
   REGION "BUTTON SELECTION BUTTONS"
       FOR #i := 0 TO "BUTTON_COUNT" DO
           #t_interface.buttons[#i].animate := "Bool.Animate"(true_color := "GREEN_LIGHT_BACKGROUND",
                                                              false_color := "GRAY_BACKGROUND",
                                                              evaluation_signal := #interface.buttons[#i].actuate);
           #t_interface.buttons[#i].enable := TRUE;
           #t_interface.buttons[#i].visible := TRUE;
           IF #selected.btns[#i] THEN
               #t_interface.buttons[#i].animate := "BLUE_LIGHT_BACKGROUND";
           END_IF;
       END_FOR;
   END_REGION


   REGION "DRAW"
       #interface := #t_interface;
   END_REGION
END_FUNCTION

FUNCTION "Pop Up: Select Buttons: Pulse Ints to Bools" : Void   // FC118, SCL
{ S7_Optimized_Access := 'TRUE' }
VERSION : 0.1
   VAR_INPUT
      pulses_as_ints : Array[0.."BUTTON_COUNT"] of Int;
   END_VAR
   VAR_OUTPUT
      pulses_as_bools : Array[0.."BUTTON_COUNT"] of Bool;
   END_VAR
   VAR_TEMP
      i : Int;
      ret : Array[0.."BUTTON_COUNT"] of Bool;
   END_VAR
BEGIN
   REGION "MAP TO BOOLS"
       FOR #i := 0 TO "BUTTON_COUNT" DO
           #ret[#i] := #pulses_as_ints[#i].%X0;
       END_FOR;
   END_REGION

   REGION "RETURN"
       #pulses_as_bools := #ret;
   END_REGION
END_FUNCTION

// folder: Display: Warehouse/Pop Ups/Select Station

FUNCTION_BLOCK "Pop Up: Select Stations"   // FB21, SCL
{ S7_Optimized_Access := 'TRUE' }
VERSION : 0.1
   VAR_INPUT
      all_stations : "Station: All Stations";
      saved_WIPs : "Recipe: HMI Stations Saved Wips";
   END_VAR
   VAR_IN_OUT
      interface : "Select Station";
      meta_data : "Setting Meta Data";
   END_VAR
   VAR
      "inst Patch for Table Nav in Select Station Popup" : "Patch for Table Nav in Select Station Popup";
      "inst Select Station Button Pulses" : "Pulses: Button Collection";
      "inst Selection Change" : "Selected_Stations.Selection_Change";
      "inst Table Nav" : "Table Nav";
      vis_stns_as_dint : Array[0.."_SELECT_STATION_BUTTON_COUNT"] of DInt;
      visable_stns : Array[0.."_SELECT_STATION_BUTTON_COUNT"] of Int;
   END_VAR
   VAR_TEMP
      actuations_as_ints : Array[0.."_SELECT_STATION_BUTTON_COUNT"] of Int;
      actuation_pulses : Array[0.."_SELECT_STATION_BUTTON_COUNT"] of Bool;
      actuation_pulses_as_int : Array[0.."_SELECT_STATION_BUTTON_COUNT"] of Int;
      blank_station : "Station: Single Station";
      i : Int;
      nav_pulses : Int;
      p_stn : DInt;
      selectable_stns_as_dint : Array[0.."STATION_COUNT"] of DInt;
      t_selection_change : "Station Selection Change";
   END_VAR
   // visable_stns[0] := 0;
   // visable_stns[1] := 1;
   // visable_stns[2] := 2;
   // visable_stns[3] := 3;
   // visable_stns[4] := 4;
   // visable_stns[5] := 5;
   // visable_stns[6] := 6;
   // visable_stns[7] := 7;
   // visable_stns[8] := 8;
   // visable_stns[9] := 9;
   // visable_stns[10] := 10;
   // visable_stns[11] := 11;
BEGIN
   REGION "ANIMATIONS"
       "Pop Up: Select Stations: Animations"(all_stations := #all_stations,
                                             meta_data := #meta_data,
                                             visable_stns := #visable_stns,
                                             interface := #interface);
   END_REGION


   REGION "CLEAR SELECTION CHANGE"
       #meta_data.station_selection_change := #t_selection_change;
   END_REGION


   REGION "SELECT STATION BUTTON PULSES"
       "Pop Up: Map Select Button Actuations"(screen_elements := #interface.stn_select_btns,
                                              actuations_as_ints := #actuations_as_ints);
       #"inst Select Station Button Pulses"(btns := #actuations_as_ints,
                                            pulses := #actuation_pulses_as_int);
       "Pop Up: Select Stations: Pulse Ints to Bools"(pulses_as_ints := #actuation_pulses_as_int,
                                                      pulses_as_bools => #actuation_pulses);
   END_REGION


   REGION "PERFORM STATION SELECTION"
       FOR #i := 0 TO "_SELECT_STATION_BUTTON_COUNT" DO
           IF #visable_stns[#i] <> -1 THEN
               "Toggle"(pulse := #actuation_pulses[#i],
                        state := #meta_data.selected_stations.stns[#visable_stns[#i]]);
           END_IF;
       END_FOR;
       #meta_data.selected_stations.count := "Count Selected Stations"(#meta_data.selected_stations.stns);
   END_REGION


   REGION "SCAN FOR CHANGE TO STATION SELECTION"
       #"inst Selection Change"(selected_stns := #meta_data.#selected_stations,
                                station_change => #meta_data.station_selection_change);
   END_REGION


   REGION "BUILD SELECTABLE STATION LIST"
       IF #meta_data.station_selection_change.selection_change OR "FirstScan" THEN
           "Pop Up: Select Stations: Build Selectable Station List"(saved_wips := #saved_WIPs,
                                                                    all_stations := #all_stations,
                                                                    meta_data := #meta_data);
       END_IF;
   END_REGION


   REGION "TABLE NAV"

       // when there are more selectable stations than buttons
       IF #meta_data.selectable_stations.count > "_SELECT_STATION_BUTTON_COUNT" THEN
           #"inst Table Nav"(first_null_index := #meta_data.selectable_stations.count,
                             tblData := #selectable_stns_as_dint,
                             tblDisp := #vis_stns_as_dint,
                             tableNav := #interface.nav_bar.plc,
                             rowIndices := #vis_stns_as_dint);
           // patch for table nav to work with selectable stations
           #"inst Patch for Table Nav in Select Station Popup"(nav_bar := #interface.nav_bar.plc,
                                                               meta_data := #meta_data,
                                                               vis_stns_as_dint := #vis_stns_as_dint,
                                                               visable_stns := #visable_stns);
       END_IF;

       // when there are fewer selectable stations than buttons
       IF #meta_data.selectable_stations.count <= "_SELECT_STATION_BUTTON_COUNT" + 1 THEN
           IF #meta_data.station_selection_change.selection_change THEN
               "Array.Int.Fill"(value:="NULL_TOKEN",
                                int_array := #visable_stns);
               FOR #i := 0 TO #meta_data.selectable_stations.count - 1 DO
                   #visable_stns[#i] := #meta_data.selectable_stations.stns[#i];
               END_FOR;
           END_IF;
       END_IF;


   END_REGION
END_FUNCTION_BLOCK

FUNCTION_BLOCK "Selected_Stations.Selection_Change"   // FB23, SCL
{ S7_Optimized_Access := 'TRUE' }
VERSION : 0.1
   VAR_INPUT
      selected_stns : "Selected Stations";
   END_VAR
   VAR_OUTPUT
      station_change : "Station Selection Change";
   END_VAR
   VAR
      old : Struct
         selected_stns : "Selected Stations";
      END_STRUCT;
   END_VAR
   VAR_TEMP
      i : Int;
      ret : "Station Selection Change";
   END_VAR
BEGIN
   REGION "SCAN FOR CHANGE"
       FOR #i := 0 TO "STATION_COUNT" DO
           IF #selected_stns.stns[#i] <> #old.selected_stns.stns[#i] THEN
               #ret.selection_change := TRUE;
               #ret.station_index := #i;
               IF #selected_stns.stns[#i] AND NOT #old.selected_stns.stns[#i] THEN
                   #ret.rising := TRUE;
                   #ret.falling := FALSE;
               END_IF;
               IF NOT #selected_stns.stns[#i] AND #old.selected_stns.stns[#i] THEN
                   #ret.rising := FALSE;
                   #ret.falling := TRUE;
               END_IF;
               EXIT;
           END_IF;
       END_FOR;
   END_REGION


   REGION "SAVE TO OLD"
       #old.selected_stns := #selected_stns;
   END_REGION


   REGION "RETURN"
       #station_change.falling := #ret.falling;
       #station_change.rising := #ret.rising;
       #station_change.selection_change := #ret.selection_change;
       #station_change.station_index := #ret.station_index;
   END_REGION
END_FUNCTION_BLOCK

FUNCTION_BLOCK "Patch for Table Nav in Select Station Popup"   // FB24, SCL
{ S7_Optimized_Access := 'TRUE' }
VERSION : 0.1
   VAR_INPUT
      nav_bar : "Nav Bar Data: PLC";
      meta_data : "Setting Meta Data";
   END_VAR
   VAR_IN_OUT
      vis_stns_as_dint : Array[0.."_SELECT_STATION_BUTTON_COUNT"] of DInt;
      visable_stns : Array[0.."_SELECT_STATION_BUTTON_COUNT"] of Int;
   END_VAR
   VAR
      old_nav : "Nav Bar Data: PLC";
   END_VAR
   VAR_TEMP
      first_row : Int;
      i : Int;
      nav_pulse : Bool;
      p_visable_row : Int;
      search_term : Int;
      t_visable_stns : Array[0.."_SELECT_STATION_BUTTON_COUNT"] of Int;
   END_VAR
BEGIN
   REGION "PULSE FROM ANY NAV BUTTON"
       IF NOT #old_nav.top.actuate AND #nav_bar.top.actuate THEN
           #nav_pulse := TRUE;
       END_IF;
       IF NOT #old_nav.pageUp.actuate AND #nav_bar.pageUp.actuate THEN
           #nav_pulse := TRUE;
       END_IF;
       IF NOT #old_nav.lineUp.actuate AND #nav_bar.lineUp.actuate THEN
           #nav_pulse := TRUE;
       END_IF;
       IF NOT #old_nav.lineDown.actuate AND #nav_bar.lineDown.actuate THEN
           #nav_pulse := TRUE;
       END_IF;
       IF NOT #old_nav.pageDown.actuate AND #nav_bar.pageDown.actuate THEN
           #nav_pulse := TRUE;
       END_IF;
       IF NOT #old_nav.bottom.actuate AND #nav_bar.bottom.actuate THEN
           #nav_pulse := TRUE;
       END_IF;
   END_REGION



   REGION "REMAP VISIBLE STATIONS BASED ON SELECTABLE STATIONS"

       REGION "NAV REMAP"
           IF #nav_pulse THEN
               FOR #i := 0 TO "_SELECT_STATION_BUTTON_COUNT" DO
                   #t_visable_stns[#i] := #meta_data.selectable_stations.stns[DINT_TO_INT(#vis_stns_as_dint[#i])];
                   #vis_stns_as_dint[#i] := #t_visable_stns[#i];
               END_FOR;
               #visable_stns := #t_visable_stns;
           END_IF;
       END_REGION

       REGION "SELECTION REMAP"
           IF #meta_data.station_selection_change.selection_change THEN
               #search_term := #visable_stns[0];
               #first_row := "Array.Int.Search"(array_of_int := #meta_data.selectable_stations.stns,
                                                 search_term := #search_term);
               WHILE #first_row = "NULL_TOKEN" DO
                   #search_term -= 1;
                   IF #search_term < 0 THEN
                       #search_term := 0;
                       EXIT;
                   END_IF;
                   #first_row := "Array.Int.Search"(array_of_int := #meta_data.selectable_stations.stns,
                                                     search_term := #search_term);
               END_WHILE;
               // direct write access required to keep collapsed or uncollapsed
               // format after nav button press
               "EMP IDB"."inst Pop Up: Select Station"."inst Table Nav".r1 := #first_row;
               FOR #i := 0 TO "_SELECT_STATION_BUTTON_COUNT" DO
                   #p_visable_row := #first_row + #i;
                   IF #p_visable_row >= #meta_data.selectable_stations.count THEN
                       #p_visable_row -= #meta_data.selectable_stations.count;
                   END_IF;
                   #t_visable_stns[#i] := #meta_data.selectable_stations.stns[#p_visable_row];
                   #vis_stns_as_dint[#i] := #t_visable_stns[#i];
               END_FOR;
               #visable_stns := #t_visable_stns;
           END_IF;
       END_REGION
   (*    
       IF #meta_data.selection_change.selection_change THEN

           REGION "COPY TO LOCAL"
               FOR #i := 0 TO "slct_stn_btn_count" DO
                   #t_visable_stns[#i] := DINT_TO_INT(#vis_stns_as_dint[#i]);
               END_FOR;
           END_REGION



           IF #meta_data.selection_change.falling AND #meta_data.selected_stations.count = 0 THEN
               #first_row := DINT_TO_INT(#vis_stns_as_dint[0]);
               FOR #i := 0 TO "slct_stn_btn_count" DO
                   #t_visable_stns[#i] := #first_row + #i;
                   IF #t_visable_stns[#i] > "stnCount" THEN
                       #t_visable_stns[#i] -= "stnCount" + 1;
                   END_IF;
               END_FOR;
           END_IF;

           IF #meta_data.selection_change.selection_change AND #meta_data.selected_stations.count <> 0 THEN
               FOR #i := 0 TO "slct_stn_btn_count" DO
                   IF DINT_TO_INT(#vis_stns_as_dint[#i]) > #meta_data.selectable_stations.count - 1 THEN
                       #t_visable_stns[#i] := DINT_TO_INT(#vis_stns_as_dint[#i]) - #meta_data.selectable_stations.count;
                   END_IF;
                   IF DINT_TO_INT(#vis_stns_as_dint[#i]) <= #meta_data.selectable_stations.count - 1 THEN

                   END_IF;
               END_FOR;
           END_IF;


           REGION "RETURN"
               FOR #i := 0 TO "slct_stn_btn_count" DO
                   #vis_stns_as_dint[#i] := INT_TO_DINT(#t_visable_stns[#i]);
               END_FOR;
               #visable_stns := #t_visable_stns;
           END_REGION


       END_IF;
   *)    

   END_REGION


   REGION "SAVE FOR CHANGE DETECTION"
       #old_nav := #nav_bar;
   END_REGION
END_FUNCTION_BLOCK

FUNCTION "Populate Station Name" : WString   // FC100, SCL
{ S7_Optimized_Access := 'TRUE' }
VERSION : 0.1
   VAR_INPUT
      lines : Int;
      stn : "Station: Single Station";
   END_VAR
   VAR_TEMP
      ret : WString;
      dz : WString;
   END_VAR
   VAR CONSTANT
      line_feed : WString := WSTRING#'$L';
   END_VAR
BEGIN
   REGION "FORMAT STRING"
       #dz := "Strip Sign"(USINT_TO_WSTRING(#stn.id.dropZone));
       #dz := "Add Leading"("Leading Character" := wchar#'0',
                            "Desired Length" := 2,
                            "String" := #dz);
   END_REGION

   REGION "ONE LINE"
       IF #lines = 1 THEN
           #ret := CONCAT_WSTRING(IN1 := #stn.id.lineName,
                                  IN2 := #dz);
       END_IF;
   END_REGION


   REGION "MORE THAN ONE LINE"
       IF #lines > 1 THEN
           #ret := CONCAT_WSTRING(IN1 := #stn.id.lineName,
                                  IN2 := #line_feed,
                                  IN3 := #dz);
       END_IF;
   END_REGION


   REGION "INVALID ENTRY"
       IF #lines < 1 THEN
           #ret := WString#'invalid line count';
       END_IF;
   END_REGION


   #"Populate Station Name" := #ret;
END_FUNCTION

FUNCTION "Pop Up: Select Stations: Map Select Button Acutations" : Void   // FC101, SCL
{ S7_Optimized_Access := 'TRUE' }
VERSION : 0.1
   VAR_INPUT
      select_btns : Array[0.."_SELECT_STATION_BUTTON_COUNT"] of "Push Button Data";
   END_VAR
   VAR_OUTPUT
      btn_actuations : Array[0.."_SELECT_STATION_BUTTON_COUNT"] of Int;
   END_VAR
   VAR_TEMP
      i : Int;
      ret : Array[0.."_SELECT_STATION_BUTTON_COUNT"] of Int;
   END_VAR
BEGIN
   REGION "MAP ACTUATIONS"
       FOR #i := 0 TO "_SELECT_STATION_BUTTON_COUNT" DO
           IF #select_btns[#i].actuate THEN
               #ret[#i] := 1;
           END_IF;
       END_FOR;
   END_REGION


   REGION "RETURN"
       #btn_actuations := #ret;
   END_REGION
END_FUNCTION

FUNCTION "Pop Up: Select Stations: Pulse Ints to Bools" : Void   // FC102, SCL
{ S7_Optimized_Access := 'TRUE' }
VERSION : 0.1
   VAR_INPUT
      pulses_as_ints : Array[0.."_SELECT_STATION_BUTTON_COUNT"] of Int;
   END_VAR
   VAR_OUTPUT
      pulses_as_bools : Array[0.."_SELECT_STATION_BUTTON_COUNT"] of Bool;
   END_VAR
   VAR_TEMP
      i : Int;
      ret : Array[0.."_SELECT_STATION_BUTTON_COUNT"] of Bool;
   END_VAR
BEGIN
   REGION "MAP TO BOOLS"
       FOR #i := 0 TO "_SELECT_STATION_BUTTON_COUNT" DO
           #ret[#i] := #pulses_as_ints[#i].%X0;
       END_FOR;
   END_REGION

   REGION "RETURN"
       #pulses_as_bools := #ret;
   END_REGION
END_FUNCTION

FUNCTION "Pop Up: Select Stations: Build Selectable Station List" : Void   // FC104, SCL
{ S7_Optimized_Access := 'TRUE' }
VERSION : 0.1
   VAR_INPUT
      saved_wips : "Recipe: HMI Stations Saved Wips";
      all_stations : "Station: All Stations";
   END_VAR
   VAR_IN_OUT
      meta_data : "Setting Meta Data";
   END_VAR
   VAR_TEMP
      eval_station_is_hmi : Bool;
      blank_stn : "Station: Single Station";
      i : Int;
      states : "Selectable Station States";
      md : "Setting Meta Data";
   END_VAR
   VAR CONSTANT
      initialize : String := 'initialize';
      all : String := 'all';
      non_hmi : String := 'non_hmi';
      hmi : String := 'hmi';
   END_VAR
BEGIN
   REGION "NOTES"
       (*
       The UDT containing all stations is too large to be instantiated in temp
       memory for this function. This is why you will see an initialization loop
       instead of a temp variable that gets returned later.
       *)
   END_REGION


   REGION "FOR ANY STATE"

       REGION "COPY TO LOCAL"
           #md := #meta_data;
       END_REGION

       REGION "SELECTED STATION IS HMI"
           IF #md.station_selection_change.rising THEN
               #eval_station_is_hmi := "Station.Is_HMI_Station"(#all_stations.stn[#md.station_selection_change.station_index]);
           END_IF;
           IF #md.station_selection_change.falling AND #md.selected_stations.count = 1 THEN
               #eval_station_is_hmi := "Station.Is_HMI_Station"(#all_stations.stn["Get First Selected Station"(#md.selected_stations.stns)]);
           END_IF;
       END_REGION

   END_REGION


   REGION "SET STATE"

       REGION "ALL"
           // on first scan
           IF "FirstScan" THEN
               #states := "Set Selectable Station States"(#all);
               GOTO EVAL;
           END_IF;
           // on selection change where last selected station is de-selected
           IF #md.station_selection_change.falling AND #md.selected_stations.count = 0 THEN
               #states := "Set Selectable Station States"(#all);
               GOTO EVAL;
           END_IF;
       END_REGION

       REGION "NON HMI"
           // when no stations are selected and a non-hmi station is selected
           IF #md.station_selection_change.selection_change (*AND #selected_stn_count = 1*) THEN
               IF NOT #eval_station_is_hmi THEN
                   #states := "Set Selectable Station States"(#non_hmi);
                   GOTO EVAL;
               END_IF;
           END_IF;
       END_REGION

       REGION "HMI"
           // when no stations are selected and an hmi station is selected
           IF #md.station_selection_change.selection_change (*AND #selected_stn_count = 1*) THEN
               IF #eval_station_is_hmi THEN
                   #states := "Set Selectable Station States"(#hmi);
                   GOTO EVAL;
               END_IF;
           END_IF;
       END_REGION

   END_REGION


   REGION "STATE LOGIC"
   EVAL:

       REGION "ALL"
           IF #states.all THEN
               "Array.Int.Fill"(value:="NULL_TOKEN",
                                int_array := #md.selectable_stations.stns);
               FOR #i := 0 TO "STATION_COUNT" DO
                   #md.selectable_stations.stns[#i] := #i;
               END_FOR;
               #md.selectable_stations.count := "STATION_COUNT" + 1;
               GOTO RTRN;
           END_IF;
       END_REGION


       REGION "NON-HMI"
           IF #states.non_hmi THEN
               "Array.Int.Fill"(value:="NULL_TOKEN",
                                int_array := #md.selectable_stations.stns);
               #md.selectable_stations := "Pop Up: Select Stations: Build Non-HMI List"(#all_stations);
               GOTO RTRN;
           END_IF;
       END_REGION


       REGION "HMI"
           IF #states.hmi THEN
               "Array.Int.Fill"(value:="NULL_TOKEN",
                                int_array := #md.selectable_stations.stns);
               #md.selectable_stations := "Pop Up: Select Stations: Build HMI List"(saved_wips := #saved_wips,
                                                                                    meta_data := #md);
               GOTO RTRN;
           END_IF;
       END_REGION

   END_REGION


   REGION "RETURN"
   RTRN:
       #meta_data := #md;
   END_REGION
END_FUNCTION

FUNCTION "Set Selectable Station States" : "Selectable Station States"   // FC107, SCL
{ S7_Optimized_Access := 'TRUE' }
VERSION : 0.1
   VAR_INPUT
      desired_state : String;
   END_VAR
   VAR_TEMP
      ret : "Selectable Station States";
   END_VAR
   VAR CONSTANT
      initialize : String := 'initialize';
      all : String := 'all';
      non_hmi : String := 'non_hmi';
      hmi : String := 'hmi';
   END_VAR
BEGIN
   REGION "SET ALL"
       IF #desired_state = #all THEN
           #ret.all := TRUE;
       END_IF;
   END_REGION


   REGION "SET NON_HMI"    
       IF #desired_state = #non_hmi THEN
           #ret.non_hmi := TRUE;
       END_IF;
   END_REGION


   REGION "SET HMI"
       IF #desired_state = #hmi THEN
           #ret.hmi := TRUE;
       END_IF;
   END_REGION


   REGION "RETURN"
       #"Set Selectable Station States" := #ret;
   END_REGION
END_FUNCTION

FUNCTION "Pop Up: Select Stations: Build Non-HMI List" : "Selectable Stations"   // FC110, SCL
{ S7_Optimized_Access := 'TRUE' }
VERSION : 0.1
   VAR_INPUT
      stns : "Station: All Stations";
   END_VAR
   VAR_TEMP
      i : Int;
      t_selectable_stations : "Selectable Stations";
      p_list : Int;
   END_VAR
   VAR CONSTANT
      null_value : Int := -1;
   END_VAR
BEGIN
   REGION "NOTES"
       (*
       Checks to see if the evaluation station matches each station
       in the context of being or not being an HMI station.
       Returns the list of matching stations.
       *)
   END_REGION


   REGION "INITIALIZE"
       "Array.Int.Fill"(value := "NULL_TOKEN",
                        int_array := #t_selectable_stations.stns);
   END_REGION


   REGION "BUILD LIST"
       FOR #i := 0 TO "STATION_COUNT" DO
           IF NOT "Station.Is_HMI_Station"(#stns.stn[#i]) THEN
               #t_selectable_stations.stns[#p_list] := #i;
               #p_list += 1;
           END_IF;
       END_FOR;
       #t_selectable_stations.count := #p_list;
   END_REGION


   REGION "RETURN"
       #"Pop Up: Select Stations: Build Non-HMI List" := #t_selectable_stations;
   END_REGION
END_FUNCTION

FUNCTION "Pop Up: Select Stations: Build HMI List" : "Selectable Stations"   // FC112, SCL
{ S7_Optimized_Access := 'TRUE' }
VERSION : 0.1
   VAR_INPUT
      meta_data : "Setting Meta Data";
      saved_wips : "Recipe: HMI Stations Saved Wips";
   END_VAR
   VAR_TEMP
      md : "Setting Meta Data";
      selected_stations_indices : Array[0.."STATION_COUNT"] of Int;
   END_VAR
BEGIN
   REGION "SET UP LOCALS"
       #md := #meta_data;
       "Array.Int.Fill"(value:= "NULL_TOKEN",
                        int_array:=#selected_stations_indices);
       #md.selectable_stations.count := 0;
       "Selected_Stations.Indices"(selected_stations := #md.selected_stations,
                                   selected_stations_indices := #selected_stations_indices);
   END_REGION


   REGION "SINGLE STATION"
       IF #md.selected_stations.count = 1 THEN
           "Build HMI List: Single Selected Station"(saved_wips := #saved_wips,
                                                     selected_stations_indices := #selected_stations_indices,
                                                     meta_data := #md);
       END_IF;
   END_REGION


   REGION "MULTIPLE STATIONS SELECTED"
       IF #md.selected_stations.count >= 2 THEN
           "Build HMI List: Multiple Selected Stations"(saved_wips := #saved_wips,
                                                        meta_data := #md,
                                                        selected_stations_indices := #selected_stations_indices);
       END_IF;
   END_REGION


   REGION "RETURN"
       #"Pop Up: Select Stations: Build HMI List" := #md.selectable_stations;
   END_REGION
END_FUNCTION

FUNCTION "Pop Up: Select Stations: Animations" : Void   // FC119, SCL
{ S7_Optimized_Access := 'TRUE' }
VERSION : 0.1
   VAR_INPUT
      all_stations : "Station: All Stations";
      meta_data : "Setting Meta Data";
      visable_stns : Array[0.."_SELECT_STATION_BUTTON_COUNT"] of Int;
   END_VAR
   VAR_IN_OUT
      interface : "Select Station";
   END_VAR
   VAR_TEMP
      i : Int;
      t_interface : "Select Station";
      labels : Array[0.."_SELECT_STATION_BUTTON_COUNT"] of String;
      t_selected_stns : Array[0.."STATION_COUNT"] of Int;
   END_VAR
BEGIN
   REGION "COPY TO LOCAL"
       #t_interface := #interface;
   END_REGION


   REGION "ANIMATE CLOSE SCREEN BUTTON"
       #t_interface.close_screen.animate := "Bool.Animate"(true_color := "GREEN_LIGHT_BACKGROUND",
                                                           false_color := "RED_LIGHT_BACKGROUND",
                                                           evaluation_signal := #t_interface.close_screen.actuate);
   END_REGION


   REGION "ANIMATE STATION SELECT BUTTONS"

       REGION "POPULATE STATION NAMES"
           FOR #i := 0 TO "_SELECT_STATION_BUTTON_COUNT" DO
               IF #visable_stns[#i] <> "NULL_TOKEN" THEN
                   #labels[#i] := WSTRING_TO_STRING("Populate Station Name"(lines := 2, stn := #all_stations.stn[#visable_stns[#i]]));
               END_IF;
           END_FOR;
       END_REGION

       REGION "BECAUSE MOVE BLOCK VARIANT DOESN'T SUPPORT ARRAYS OF BOOL"
           FOR #i := 0 TO "STATION_COUNT" DO
               IF #meta_data.selected_stations.stns[#i] THEN
                   #t_selected_stns[#i] := 1;
               END_IF;
           END_FOR;
       END_REGION

       REGION "ANIMATE"
           "Animate Array: PB Data"(labels := #labels,
                                    pb_data := #t_interface.stn_select_btns,
                                    selected_elements := #t_selected_stns,
                                    visible_elements := #visable_stns,
                                    visible_pb_count := #meta_data.selectable_stations.count);
       END_REGION

   END_REGION


   REGION "ANIMATE NAV BAR"
       "Pop Up: Nav Bar: Animate"(selectable_element_count := #meta_data.selectable_stations.count,
                                  visible_rows := "_SELECT_STATION_BUTTON_COUNT",
                                  nav_bar := #t_interface.nav_bar);
   END_REGION


   REGION "DRAW"
       #interface := #t_interface;
   END_REGION
END_FUNCTION

FUNCTION "Animate Array: PB Data" : Void   // FC136, SCL
{ S7_Optimized_Access := 'TRUE' }
VERSION : 0.1
   VAR_INPUT
      labels : Variant;
      pb_data : Variant;
      selected_elements : Variant;
      visible_elements : Variant;
      visible_pb_count : Int;
   END_VAR
   VAR_TEMP
      i : Int;
      len_labels : UDInt;
      len_pb_data : Struct
         as_udint : UDInt;
         as_int : Int;
      END_STRUCT;
      len_selected_elements : UDInt;
      len_visible_elements : UDInt;
      status : Int;
      t_labels : Array[0..#complex_u_bound] of String;
      t_pb_data : Array[0..#complex_u_bound] of "Push Button Data";
      t_selected_elements : Array[0..#simple_u_bound] of Int;
      t_visible_elements : Array[0..#simple_u_bound] of Int;
   END_VAR
   VAR CONSTANT
      simple_u_bound : Int := 49;
      complex_u_bound : Int := 19;
   END_VAR
BEGIN
   REGION "GET ARRAY PARAMETERS"
       #len_labels := CountOfElements(#labels);
       #len_pb_data.as_udint := CountOfElements(#pb_data);
       #len_pb_data.as_int := UDINT_TO_INT(#len_pb_data.as_udint) - 1;
       #len_selected_elements := CountOfElements(#selected_elements);
       #len_visible_elements := CountOfElements(#visible_elements);
   END_REGION


   REGION "COPY TO LOCAL"
       #status := MOVE_BLK_VARIANT(SRC := #labels,
                                   COUNT := #len_labels,
                                   SRC_INDEX := 0,
                                   DEST_INDEX := 0,
                                   DEST => #t_labels);
       #status := MOVE_BLK_VARIANT(SRC := #pb_data,
                                   COUNT := #len_pb_data.as_udint,
                                   SRC_INDEX := 0,
                                   DEST_INDEX := 0,
                                   DEST => #t_pb_data);
       #status := MOVE_BLK_VARIANT(SRC := #selected_elements,
                                   COUNT := #len_selected_elements,
                                   SRC_INDEX := 0,
                                   DEST_INDEX := 0,
                                   DEST => #t_selected_elements);
       #status := MOVE_BLK_VARIANT(SRC := #visible_elements,
                                   COUNT := #len_visible_elements,
                                   SRC_INDEX := 0,
                                   DEST_INDEX := 0,
                                   DEST => #t_visible_elements);
   END_REGION

   REGION "FOR EACH BUTTON"
       FOR #i := 0 TO #len_pb_data.as_int DO

           REGION "ENABLE"
               #t_pb_data[#i].enable := "Animate Array: PB Data Activation"(element_index := #i,
                                                                            visible_element_count := #visible_pb_count);
           END_REGION

           REGION "VISIBLITY"
               #t_pb_data[#i].visible := "Animate Array: PB Data Activation"(element_index := #i,
                                                                             visible_element_count := #visible_pb_count);
           END_REGION

           REGION "NO FURTHER OPERATIONS ON NULL VALUE"
               IF #t_visible_elements[#i] = "NULL_TOKEN" THEN
                   CONTINUE;
               END_IF;
           END_REGION

           REGION "ACTUATION: NOT SELECTED"
               IF #t_selected_elements[#t_visible_elements[#i]] = 0 THEN
                   #t_pb_data[#i].animate := "Bool.Animate"(true_color := "GREEN_LIGHT_BACKGROUND",
                                                            false_color := "GRAY_BACKGROUND",
                                                            evaluation_signal := #t_pb_data[#i].actuate);
               END_IF;
           END_REGION

           REGION "ACTUATION: SELECTED"
               IF #t_selected_elements[#t_visible_elements[#i]] = 1 THEN
                   #t_pb_data[#i].animate := "Bool.Animate"(true_color := "GREEN_LIGHT_BACKGROUND",
                                                            false_color := "BLUE_LIGHT_BACKGROUND",
                                                            evaluation_signal := #t_pb_data[#i].actuate);
               END_IF;
           END_REGION

           REGION "LABEL"
               #t_pb_data[#i].label := STRING_TO_WSTRING(#t_labels[#i]);
           END_REGION

       END_FOR;
   END_REGION


   REGION "DRAW"
       #status := MOVE_BLK_VARIANT(SRC := #t_pb_data,
                                   COUNT := #len_pb_data.as_udint,
                                   SRC_INDEX := 0,
                                   DEST_INDEX := 0,
                                   DEST => #pb_data);
   END_REGION
END_FUNCTION

FUNCTION "Build HMI List: Single Selected Station" : Void   // FC146, SCL
{ S7_Optimized_Access := 'TRUE' }
VERSION : 0.1
   VAR_INPUT
      saved_wips : "Recipe: HMI Stations Saved Wips";
      selected_stations_indices : Array[0.."STATION_COUNT"] of Int;
   END_VAR
   VAR_IN_OUT
      meta_data : "Setting Meta Data";
   END_VAR
   VAR_TEMP
      station : "WIP: Station";
      has_matching_wip : Bool;
      i : Int;
      j : Int;
   END_VAR
BEGIN
   REGION "GET SELECTED STATION"
       #station := "WIP.Global_Index_to_Station"(index := #selected_stations_indices[0],
                                                     wip_stations := #saved_wips);
   END_REGION

   REGION "SELF IS ALWAYS SELECTABLE"
       #meta_data.selectable_stations.stns[#meta_data.selectable_stations.count] := #station.pStn;
       #meta_data.selectable_stations.count += 1;
   END_REGION

   REGION "CHECK STATIONS FOR MATCHING WIPS"
       FOR #j := 0 TO "HMI_STATION_COUNT" DO

           REGION "DONT RUN IF SELECTED AND EVALUATION STATIONS MATCH"
               IF #station.pStn = #saved_wips.stn[#j].pStn THEN
                   CONTINUE;
               END_IF;
           END_REGION

           REGION "ADD TO LIST ON MATCHING WIP"
               #has_matching_wip := "Array.DInt.Intersect_Exists"(a := #station.wip,
                                                                    b := #saved_wips.stn[#j].wip,
                                                                    null_value := "NULL_TOKEN");
               IF #has_matching_wip THEN
                   #meta_data.selectable_stations.stns[#meta_data.selectable_stations.count] := #saved_wips.stn[#j].pStn;
                   #meta_data.selectable_stations.count += 1;
               END_IF;
           END_REGION

       END_FOR;
   END_REGION
END_FUNCTION

FUNCTION "Build HMI List: Multiple Selected Stations" : Void   // FC147, SCL
{ S7_Optimized_Access := 'TRUE' }
VERSION : 0.1
   VAR_INPUT
      saved_wips : "Recipe: HMI Stations Saved Wips";
   END_VAR
   VAR_IN_OUT
      meta_data : "Setting Meta Data";
      selected_stations_indices : Array[0.."STATION_COUNT"] of Int;
   END_VAR
   VAR_TEMP
      selected_station_a_WIP_codes : "Selectable Wips";
      selected_station_b_WIP_codes : "Selectable Wips";
      intersect_of_WIPs : Array[0.."WIP_COUNT"] of DInt;
      has_matching_wip : Bool;
      i : Int;
   END_VAR
BEGIN
   REGION "SELECTED STATIONS ARE ALWAYS SELECTABLE"
       FOR #i := 0 TO #meta_data.selected_stations.count DO
           #meta_data.selectable_stations.stns[#i] := #selected_stations_indices[#i];
       END_FOR;
   END_REGION

   REGION "MAP SELECTED STATIONS TO ARRAY OF INDICIES"
       "Map Selected Stations to Int Array"(selected_stations := #meta_data.selected_stations,
                                            selected_stations_indicies => #selected_stations_indices);
   END_REGION

   REGION "GET FIRST TWO SELECTED STATION WIPS, SAVE AS DINT ARRAY"
       "Map WIP Codes to DInt Array"(station := "WIP.Global_Index_to_Station"(index := #selected_stations_indices[0], wip_stations := #saved_wips),
                                     WIP_array := #selected_station_a_WIP_codes.wips);
       "Map WIP Codes to DInt Array"(station := "WIP.Global_Index_to_Station"(index := #selected_stations_indices[1], wip_stations := #saved_wips),
                                     WIP_array := #selected_station_b_WIP_codes.wips);
   END_REGION

   REGION "FIND INTERSECT OF FIRST AND SECOND STATIONS WIPS" 
       "Array.DInt.Intersect"(a := #selected_station_a_WIP_codes.wips,
                                b := #selected_station_b_WIP_codes.wips,
                                null_value := INT_TO_DINT("NULL_TOKEN"),
                                intersect_array => #intersect_of_WIPs);
   END_REGION

   REGION "IF MORE THAN 2 STATIONS SELECTABLE"
       #meta_data.selectable_stations.count := "Array.Int.Count"(null_value := "NULL_TOKEN", array := #meta_data.selectable_stations.stns);
       IF #meta_data.selectable_stations.count > 2 THEN

           REGION "COMPARE SUBSIQENT STATIONS AND UPDATE SELECTABLE STATIONS"
               FOR #i := 0 TO "HMI_STATION_COUNT" DO
                   // dont evaluate selected stations
                   IF #selected_stations_indices[#i] = #meta_data.selectable_stations.stns[#i] THEN
                       CONTINUE;
                   END_IF;
                   // get wip codes of station to evaluate
                   "Map WIP Codes to DInt Array"(station := "WIP.Global_Index_to_Station"(index := #meta_data.selectable_stations.stns[#i], wip_stations := #saved_wips),
                                                 WIP_array := #selected_station_b_WIP_codes.wips);
                   // check evaluation station's wip codes against intersect array
                   #has_matching_wip := "Array.DInt.Intersect_Exists"(a := #intersect_of_WIPs,
                                                                        b := #selected_station_b_WIP_codes,
                                                                        "null_value" := "NULL_TOKEN");
                   IF #has_matching_wip THEN
                       // add to selectable 
                       #meta_data.selectable_stations.stns[#meta_data.selectable_stations.count] := #saved_wips.stn[#i].pStn;
                       #meta_data.selectable_stations.count += 1;
                       // get new intersect array
                       "Array.DInt.Intersect"(a := #intersect_of_WIPs,
                                                b := #selected_station_b_WIP_codes,
                                                null_value := "NULL_TOKEN",
                                                intersect_array => #intersect_of_WIPs);
                   END_IF;
               END_FOR;
           END_REGION

       END_IF;
   END_REGION
END_FUNCTION

// folder: Display: Warehouse/Pop Ups/Select WIP

FUNCTION_BLOCK "Pop Up: Select WIPs"   // FB28, SCL
{ S7_Optimized_Access := 'TRUE' }
VERSION : 0.1
   VAR_INPUT
      stations : "Station: All Stations";
      saved_WIPs : "Recipe: HMI Stations Saved Wips";
      wip_library : "Recipe: Wip Text Library";
   END_VAR
   VAR_IN_OUT
      interface : "Select WIP";
      meta_data : "Setting Meta Data";
   END_VAR
   VAR
      "inst Table Nav" : "Table Nav";
      "inst WIP Select Button Pulses" : "Pulses: Button Collection";
      t_selected_WIPs_as_Bools : Array[0.."WIP_COUNT"] of Bool;
      visable_WIPs : Array[0.."WIP_POPUP_BUTTON_COUNT"] of DInt;
      visable_WIPs_indices : Array[0.."WIP_POPUP_BUTTON_COUNT"] of DInt;
   END_VAR
   VAR_TEMP
      actuations_as_ints : Array[0.."WIP_POPUP_BUTTON_COUNT"] of Int;
      actuation_pulses_as_ints : Array[0.."WIP_POPUP_BUTTON_COUNT"] of Int;
      i : Int;
      indices_as_ints : Array[0.."WIP_POPUP_BUTTON_COUNT"] of Int;
      t_interface : "Select WIP";
   END_VAR
   VAR CONSTANT
      null_value : Int := -1;
   END_VAR
BEGIN
   REGION "ANIMATION"
       REGION "CONVERT DINT TO INT FOR MOVE BLOCK VARIANT"
           FOR #i := 0 TO "WIP_POPUP_BUTTON_COUNT" DO
               #indices_as_ints[#i] := DINT_TO_INT(#visable_WIPs_indices[#i]);
           END_FOR;
       END_REGION
       "Pop Up: Select WIPs: Animations"(selectable_WIP_count := #meta_data.selectable_wips.count,
                                         visable_WIPs := #visable_WIPs,
                                         selected_WIPs := #t_selected_WIPs_as_Bools,
                                         visable_WIPs_indices := #indices_as_ints,
                                         wip_library := #wip_library,
                                         interface := #interface);
   END_REGION


   REGION "SELECT WIP BUTTON PULSES"
       "Pop Up: Map Select Button Actuations"(screen_elements := #interface.select_wip_buttons,
                                              actuations_as_ints := #actuations_as_ints);
       #"inst WIP Select Button Pulses"(btns := #actuations_as_ints,
                                        pulses := #actuation_pulses_as_ints);
   END_REGION


   REGION "PERFORM WIP SELECTION"
       "Pop Up: Select WIPs: Perform Selection"(indices := #visable_WIPs_indices,
                                                pulses := #actuation_pulses_as_ints,
                                                visable_WIPs:=#visable_WIPs,
                                                selected_wips_as_bools := #t_selected_WIPs_as_Bools);
   END_REGION


   REGION "MAP SELECTION TO META DATA"
       "Pop Up: Select WIPs: Map to Meta"(actuation_pulses_as_ints := #actuation_pulses_as_ints,
                                          indices := #visable_WIPs_indices,
                                          selected_wips_as_bools := #t_selected_WIPs_as_Bools,
                                          selectable_wips := #meta_data.selectable_wips,
                                          selected_wips := #meta_data.selected_wips);
   END_REGION    


   REGION "HOUSE KEEPING FOR STATION SELECTION CHANGE"
       IF #meta_data.station_selection_change.selection_change THEN
           "Array.DInt.Fill"(int_in := INT_TO_DINT("NULL_TOKEN"),
                             array_out => #visable_WIPs);
           FOR #i := 0 TO "WIP_COUNT" DO
               #t_selected_WIPs_as_Bools[#i] := FALSE;
           END_FOR;
           "Clear WIP Selection Meta Data"(#meta_data.selected_wips);
       END_IF;
   END_REGION


   REGION "BUILD SELECTABLE WIP LIST"
       IF #meta_data.station_selection_change.selection_change THEN
           IF "Station.Is_HMI_Station"(#stations.stn[#meta_data.station_selection_change.station_index]) THEN
               "Pop Up: Select WIPs: Build Selectable List"(saved_WIPs := #saved_WIPs,
                                                            meta_data := #meta_data,
                                                            stations := #stations);
           END_IF;
       END_IF;
   END_REGION


   REGION "SHOW ALL WIPS WHEN FEWER SELECTABLE WIPS THAN BUTTONS"
       IF #meta_data.station_selection_change.selection_change AND #meta_data.selectable_wips.count - 1 <= "WIP_POPUP_BUTTON_COUNT" THEN
           "Array.DInt.Fill"(int_in := INT_TO_DINT("NULL_TOKEN"),
                             array_out => #visable_WIPs_indices);
           FOR #i := 0 TO #meta_data.selectable_wips.count - 1 DO
               #visable_WIPs[#i] := #meta_data.selectable_wips.wips[#i];
               #visable_WIPs_indices[#i] := #i;
           END_FOR;
       END_IF;
   END_REGION



   REGION "NAVIGATE THROUGH TABLE WHEN MORE SELECTABLE WIPS THAN BUTTONS"
       IF #meta_data.selectable_wips.count - 1 > "WIP_POPUP_BUTTON_COUNT" THEN

           REGION "TABLE NAVIGATION"
               #"inst Table Nav"(first_null_index := #meta_data.selectable_wips.count,
                                 tblData := #meta_data.selectable_wips.wips,
                                 tblDisp := #visable_WIPs,
                                 tableNav := #interface.nav_bar.plc,
                                 rowIndices := #visable_WIPs_indices);
           END_REGION

           REGION "MAP INDICES ON SCANS WHEN SELECTION HASN'T CHANGED"
               IF NOT #meta_data.station_selection_change.selection_change THEN
                   FOR #i := 0 TO "WIP_POPUP_BUTTON_COUNT" DO
                       #visable_WIPs[#i] := #meta_data.selectable_wips.wips[#visable_WIPs_indices[#i]];
                   END_FOR;
               END_IF;
           END_REGION

           REGION "REMAP INDICES TO TOP WHEN SELECTION HAS CHANGED"
               IF #meta_data.station_selection_change.selection_change THEN
                   FOR #i := 0 TO "WIP_POPUP_BUTTON_COUNT" DO
                       #visable_WIPs[#i] := INT_TO_DINT(#i);
                       #visable_WIPs_indices[#i] := INT_TO_DINT(#i);
                   END_FOR;
               END_IF;
           END_REGION

       END_IF;
   END_REGION
END_FUNCTION_BLOCK

FUNCTION "Pop Up: Select WIPs: Get Matching WIPs" : Void   // FC125, SCL
{ S7_Optimized_Access := 'TRUE' }
VERSION : 0.1
   VAR_INPUT
      selectable_wips : "Selectable Wips";
      station_wips : "Selectable Wips";
   END_VAR
   VAR_IN_OUT
      matching_wips : "Selectable Wips";
   END_VAR
   VAR_TEMP
      i : Int;
      j : Int;
      t_matching_wips : "Selectable Wips";
   END_VAR
BEGIN
   REGION "COPY TO LOCAL"
       "Array.DInt.Fill"(int_in := INT_TO_DINT("NULL_TOKEN"),
                         array_out => #t_matching_wips.wips);
       #t_matching_wips.count := 0;
   END_REGION

   REGION "COMPARE EACH WIP CODE IN OUTER LIST ..." 
       FOR #i := 0 TO "WIP_COUNT" DO

           REGION "LEAVE LOOP ON FIRST NULL"
               IF #selectable_wips.wips[#i] = "NULL_TOKEN" THEN
                   EXIT;
               END_IF;
           END_REGION

           REGION "WITH EACH IN INNER LIST AND ..."
               FOR #j := 0 TO "WIP_COUNT" DO

                   REGION "LEAVE LOOP ON FIRST NULL"
                       IF #station_wips.wips[#j] = "NULL_TOKEN" THEN
                           EXIT;
                       END_IF;
                   END_REGION

                   REGION "COPY MATCHES"
                       IF #selectable_wips.wips[#i] = #station_wips.wips[#j] THEN
                           #t_matching_wips.wips[#t_matching_wips.count] := #selectable_wips.wips[#i];
                           #t_matching_wips.count += 1;
                       END_IF;
                   END_REGION

               END_FOR;
           END_REGION

       END_FOR;
   END_REGION


   REGION "RETURN"
       #matching_wips := #t_matching_wips;
   END_REGION
END_FUNCTION

FUNCTION "Pop Up: Select WIPs: Build Selectable List" : Void   // FC128, SCL
{ S7_Optimized_Access := 'TRUE' }
VERSION : 0.1
   VAR_INPUT
      stations : "Station: All Stations";
      saved_WIPs : "Recipe: HMI Stations Saved Wips";
   END_VAR
   VAR_IN_OUT
      meta_data : "Setting Meta Data";
   END_VAR
   VAR_TEMP
      wip_index : Int;
      p_outer : Int;
      p_inner : Int;
      t_selectable_WIPs : "Selectable Wips";
      selected_station_WIPs : "Selected Wips";
   END_VAR
BEGIN
   REGION "NO STATIONS SELECTED"
       IF #meta_data.selected_stations.count = 0 THEN
           "Array.DInt.Fill"(int_in := INT_TO_DINT("NULL_TOKEN"),
                             array_out => #t_selectable_WIPs.wips);
           #t_selectable_WIPs.count := 0;
           GOTO RTRN;
       END_IF;
   END_REGION


   REGION "SINGLE STATION SELECTION"
       IF #meta_data.selected_stations.count = 1 THEN
           "Array.DInt.Fill"(int_in := -1,
                             array_out => #t_selectable_WIPs.wips);
           #t_selectable_WIPs.count := 0;
           #wip_index := "WIP.Global_Index_to_HMI_Station_Index"(global_index := "Get First Selected Station"(#meta_data.selected_stations.stns),
                                                                 saved_WIPs := #saved_WIPs);
           "Pop Up: Select WIPs: Map WIP Codes"(wip_station := #saved_WIPs.stn[#wip_index],
                                                selectable_wips := #t_selectable_WIPs);
           GOTO RTRN;
       END_IF;
   END_REGION


   REGION "MULTI STATION SELECTION"

       REGION "CHECK MATCHING: SELECTABLE & NEW STATION"
           #t_selectable_WIPs.wips := #meta_data.selectable_wips.wips;
           "Array.DInt.Fill"(int_in := INT_TO_DINT("NULL_TOKEN"),
                             array_out => #selected_station_WIPs.wips);
           "Map WIP Codes to DInt Array"(station := "WIP.Global_Index_to_Station"(index := #meta_data.station_selection_change.station_index, wip_stations := #saved_WIPs),
                                         WIP_array := #selected_station_WIPs.wips);
           "Pop Up: Select WIPs: Get Matching WIPs"(selectable_wips := #meta_data.selectable_wips,
                                                    station_wips := #selected_station_WIPs,
                                                    matching_wips := #t_selectable_WIPs);
       END_REGION


   END_REGION


   REGION "RETURN"
   RTRN:
       #meta_data.selectable_wips := #t_selectable_WIPs;
   END_REGION
END_FUNCTION

FUNCTION "Pop Up: Select WIPs: Map WIP Codes" : Void   // FC129, SCL
{ S7_Optimized_Access := 'TRUE' }
VERSION : 0.1
   VAR_INPUT
      wip_station : "WIP: Station";
   END_VAR
   VAR_IN_OUT
      selectable_wips : "Selectable Wips";
   END_VAR
   VAR_TEMP
      i : Int;
      t_selectable_wips : "Selectable Wips";
   END_VAR
BEGIN
   REGION "COPY TO LOCAL"
       #t_selectable_wips := #selectable_wips;
   END_REGION


   REGION "MAP VALUES"
       "Map WIP Codes to DInt Array"(station := #wip_station,
                                     WIP_array := #t_selectable_wips.wips);
   END_REGION


   REGION "COUNT SELECTABLE WIPS"
       #t_selectable_wips.count := "Count Collapsed DInt Array"(null_value := INT_TO_DINT("NULL_TOKEN"),
                                                                array := #t_selectable_wips.wips);
   END_REGION


   REGION "RETURN"
       #selectable_wips := #t_selectable_wips;
   END_REGION
END_FUNCTION

FUNCTION "Pop Up: Select WIPs: Animations" : Void   // FC134, SCL
{ S7_Optimized_Access := 'TRUE' }
VERSION : 0.1
   VAR_INPUT
      selectable_WIP_count : Int;
      selected_WIPs : Array[0.."WIP_COUNT"] of Bool;
      visable_WIPs : Array[0.."WIP_POPUP_BUTTON_COUNT"] of DInt;
      visable_WIPs_indices : Array[0.."WIP_POPUP_BUTTON_COUNT"] of Int;
      wip_library : "Recipe: Wip Text Library";
   END_VAR
   VAR_IN_OUT
      interface : "Select WIP";
   END_VAR
   VAR_TEMP
      i : Int;
      labels : Array[0.."WIP_POPUP_BUTTON_COUNT"] of String;
      t_interface : "Select WIP";
      t_selected_WIPs : Array[0.."WIP_COUNT"] of Int;
      visable_WIP_count : Int;
   END_VAR
BEGIN
   REGION "COPY TO LOCAL"
       #t_interface := #interface;
   END_REGION


   REGION "ANIMATE CLOSE SCREEN BUTTON"
       #t_interface.close_screen.animate := "Bool.Animate"(true_color := "GREEN_LIGHT_BACKGROUND",
                                                           false_color := "RED_LIGHT_BACKGROUND",
                                                           evaluation_signal := #t_interface.close_screen.actuate);
   END_REGION


   REGION "ANIMATE WIP SELECT BUTTONS" 

       REGION "WIP LABELS"
           FOR #i := 0 TO "WIP_POPUP_BUTTON_COUNT" DO
               #labels[#i] := WSTRING_TO_STRING("WIP.Code_to_WString"(wipTxtLib := #wip_library, code := #visable_WIPs[#i]));
           END_FOR;
       END_REGION

       REGION "CONVERT BOOLS TO INT FOR MOVE BLOCK VARIANT"
           FOR #i := 0 TO "WIP_COUNT" DO
               #t_selected_WIPs[#i].%X0 := #selected_WIPs[#i];
           END_FOR;
       END_REGION

